(* Logix 5000 project; controller PLC_MCC1300_75F1 vendor 1 type 14 code 166 rev 32.11; software revision 32.04; part 69 of 83 *)
(* tags used below, declared in another part *)
   CM_LineToConveyorStacker_JS1 : CM_LineToConveyorStacker;
   GP_ScadaPlate : GP_ScadaPlate;
   M317 : MAC_Conveyor_Single;
   M317_ALM : MAC_Conveyor_ALM;
   M317_Data : UDT_Convoy_SL;
   M317_HMR : MAC_Conveyor_HMR;
   M317_HMW : MAC_Conveyor_HMW;
   M317_SpaceConv_Utilities : SpaceConv_Utilities;
   M317_TON_FrontSquarLeft_timeout : TIMER;
   M317_TON_FrontSquarRight_timeout : TIMER;
   M317_TON_LatSquarLeft_timeout : TIMER;
   M317_TON_LatSquarRight_timeout : TIMER;
   M317_TON_Synchro_timeout : TIMER;
   M317_xFrontLeftTimeout : BOOL;
   M317_xFrontRightTimeout : BOOL;
   M317_xLatLeftTimeout : BOOL;
   M317_xLatRightTimeout : BOOL;
   M317_xSensorTimeout : BOOL;
   M350Popup : MAC_Popup_ZC;
   M350Popup_ALM : MAC_Popup_ZC_ALM;
   M350Popup_HMR : MAC_Popup_ZC_HMR;
   M350Popup_HMW : MAC_Popup_ZC_HMW;
   O : INT[128];
   TMP_dHalfConveyorLength : DINT;
   TMP_xEnableZoneCleaning : BOOL;
   xAlwaysOFF : BOOL;
   xAlwaysON : BOOL;
   Z300_Conveyor : UDT_StandConv[29];
   Z300_LineTracking : UDT_LINE_TRACKING;
   Z301 : MAC_Zone_ML;
   Z402 : MAC_Zone;
   Z402_HMI_rgtPlateScada_Internal : HMI_LiteData[5,2,7];
(* MainProgram, continued *)

   // Command descent frontal squaring
   103: XIC(M317.ST_xManualMode)XIC(M317_HMW.rgxMan.17)XIC(M317.OUTPUT_xDescentSquaring_1)OTE(M317_HMR.rgxMan.17);
   // Commando conveyor M317 and conveyor stacker forward
   104: XIC(M317_HMW.rgxMan.25)XIC(M317.OUTPUT_xRun_M1)XIC(CM_LineToConveyorStacker_JS1.xManualCommandFwd)OTE(M317_HMR.rgxMan.25);
   // Commando conveyor M317 and conveyor stacker backward
   105: XIC(M317_HMW.rgxMan.26)XIC(M317.OUTPUT_xReverse_M1)XIC(CM_LineToConveyorStacker_JS1.xManualCommandBkw)OTE(M317_HMR.rgxMan.26);
   // Cleaning Enabled {x|x|x|x|O}
   106: XIC(M317.ST_xCleaningAccepted)[XIC(Z402.ST_xCleaningAccepted) ,XIO(TMP_xEnableZoneCleaning) ]OTE(M317_HMR.xCleaningEnabled);
   // Virtual door Enabled {x|x|x|x|O}
   107: XIC(M317.ST_xVirtualDoorEnabled)OTE(M317_HMR.xVirtualDoorEnabled);
   // Id plate presence
   108: XIC(M317.ST_xIdPlatePresence)OTE(M317_HMR.xIdPlatePresence);
   // Machine state M1
   109: XIC(xAlwaysON)[MOV(1,M317_HMR.dState1) ,XIC(M317.OUTPUT_xRun_M1) MOV(3,M317_HMR.dState1) ,XIC(M317.OUTPUT_xReverse_M1) MOV(4,M317_HMR.dState1) ,XIC(M317.ST_xMachineAlarm) MOV(7,M317_HMR.dState1) ];
   // Machine state M2
   110: XIC(xAlwaysON)[MOV(1,M317_HMR.dState2) ,XIC(M317.OUTPUT_xRun_M2) MOV(3,M317_HMR.dState2) ,XIC(M317.OUTPUT_xReverse_M2) MOV(4,M317_HMR.dState2) ,XIC(M317.ST_xMachineAlarm) MOV(7,M317_HMR.dState2) ];
   // Machine state M3
   111: XIC(xAlwaysON)[MOV(1,M317_HMR.dState3) ,XIC(M317.OUTPUT_xRun_M3) MOV(3,M317_HMR.dState3) ,XIC(M317.OUTPUT_xReverse_M3) MOV(4,M317_HMR.dState3) ,XIC(M317.ST_xMachineAlarm) MOV(7,M317_HMR.dState3) ];
   // Machine state M4
   112: XIC(xAlwaysON)[MOV(1,M317_HMR.dState4) ,XIC(M317.OUTPUT_xRun_M4) MOV(3,M317_HMR.dState4) ,XIC(M317.OUTPUT_xReverse_M4) MOV(4,M317_HMR.dState4) ,XIC(M317.ST_xMachineAlarm) MOV(7,M317_HMR.dState4) ];
   113: XIC(M317_SpaceConv_Utilities.O_xPlateSynchronized)OTE(M317.ST_xPlateSynchronized);
   114: XIC(M317.INPUT_xSyncroPhotocell_1)XIO(M317.ST_xIdPlatePresence)XIO(M317.ST_xPlatePresence)[TON(M317_TON_Synchro_timeout,?,?) ,[XIC(M317_TON_Synchro_timeout.DN) ,XIC(M317_xSensorTimeout) ] XIC(M317.INPUT_xSyncroPhotocell_1) OTE(M317_xSensorTimeout) ];
   115: XIC(M317.INPUT_xSquaringPhotocell_1)XIO(M317.ST_xIdPlatePresence)XIO(M317.ST_xPlatePresence)[TON(M317_TON_FrontSquarRight_timeout,?,?) ,[XIC(M317_TON_FrontSquarRight_timeout.DN) ,XIC(M317_xFrontRightTimeout) ] XIC(M317.INPUT_xSquaringPhotocell_1) OTE(M317_xFrontRightTimeout) ];
   116: XIC(M317.INPUT_xSquaringPhotocell_2)XIO(M317.ST_xIdPlatePresence)XIO(M317.ST_xPlatePresence)[TON(M317_TON_FrontSquarLeft_timeout,?,?) ,[XIC(M317_TON_FrontSquarLeft_timeout.DN) ,XIC(M317_xFrontLeftTimeout) ] XIC(M317.INPUT_xSquaringPhotocell_2) OTE(M317_xFrontLeftTimeout) ];
   117: XIC(M317.INPUT_xSquaringPhotocell_3)XIO(M317.ST_xIdPlatePresence)XIO(M317.ST_xPlatePresence)[TON(M317_TON_LatSquarRight_timeout,?,?) ,[XIC(M317_TON_LatSquarRight_timeout.DN) ,XIC(M317_xLatRightTimeout) ] XIC(M317.INPUT_xSquaringPhotocell_3) OTE(M317_xLatRightTimeout) ];
   118: XIC(M317.INPUT_xSquaringPhotocell_4)XIO(M317.ST_xIdPlatePresence)XIO(M317.ST_xPlatePresence)[TON(M317_TON_LatSquarLeft_timeout,?,?) ,[XIC(M317_TON_LatSquarLeft_timeout.DN) ,XIC(M317_xLatLeftTimeout) ] XIC(M317.INPUT_xSquaringPhotocell_4) OTE(M317_xLatLeftTimeout) ];
   // State Sensor
   119: XIC(xAlwaysON)[MOV(1,M317_HMR.dStateSensor5) ,XIC(M317_xSensorTimeout) MOV(7,M317_HMR.dStateSensor5) ];
   // State Sensor
   120: XIC(xAlwaysON)[MOV(1,M317_HMR.dStateSensor3) ,[XIC(M317_ALM.rgxStoppingFault[0].2) ,XIC(M317_ALM.rgxStoppingFault[0].3) ,XIC(M317_ALM.rgxWarning[0].25) ,XIC(M317_xFrontRightTimeout) ] MOV(7,M317_HMR.dStateSensor3) ];
   // State Sensor
   121: XIC(xAlwaysON)[MOV(1,M317_HMR.dStateSensor4) ,[XIC(M317_ALM.rgxStoppingFault[0].10) ,XIC(M317_ALM.rgxStoppingFault[0].11) ,XIC(M317_ALM.rgxWarning[0].25) ,XIC(M317_xFrontLeftTimeout) ] MOV(7,M317_HMR.dStateSensor4) ];
   // State Sensor
   122: XIC(xAlwaysON)[MOV(1,M317_HMR.dStateSensor1) ,[XIC(M317_ALM.rgxWarning[0].26) ,XIC(M317_xLatRightTimeout) ] MOV(7,M317_HMR.dStateSensor1) ];
   // State Sensor
   123: XIC(xAlwaysON)[MOV(1,M317_HMR.dStateSensor2) ,[XIC(M317_ALM.rgxWarning[0].26) ,XIC(M317_xLatLeftTimeout) ] MOV(7,M317_HMR.dStateSensor2) ];
   124: XIC(M317.ST_xIdPlatePresence)GP_ScadaPlate(GP_ScadaPlate,M317_Data,6,M317_SpaceConv_Utilities.O_dHeadPosition_cmm,M317_SpaceConv_Utilities.CONST_dConveyorWidth_cmm,M317_SpaceConv_Utilities.CONST_dConveyorLength_cmm,M317_SpaceConv_Utilities.ST_xLastModLoadBkw,M317_SpaceConv_Utilities.ST_xLastModUnloadBkw,1,0,Z402_HMI_rgtPlateScada_Internal);
END_ROUTINE

ROUTINE M350Popup_Faults   (* ladder *)
   // Reset faults
   0: XIC(Z301.ST_xAlarmOff)FLL(0,M350Popup_ALM,1);
   1: XIC(M350Popup.ST_xEnableControlError)[[XIC(M350Popup.OUTPUT_xPopupLifting) XIO(M350Popup.INPUT_xPopupHigh) ,XIO(M350Popup.OUTPUT_xPopupLifting) XIO(M350Popup.INPUT_xPopupLow) ,XIO(M350Popup.INPUT_xPopupHigh) XIO(M350Popup.INPUT_xPopupLow) ] XIO(M350Popup_ALM.rgxStoppingFault[0].0) TON(M350Popup.tmON_LiftingTimeOut,?,?) ,[XIC(M350Popup.tmON_LiftingTimeOut.DN) ,XIC(M350Popup.INPUT_xPopupHigh) XIC(M350Popup.INPUT_xPopupLow) ] OTL(M350Popup_ALM.rgxStoppingFault[0].0) ];
   2: XIC(xAlwaysOFF)XIC(M350Popup.ST_xEnableControlError)XIO(M350Popup.INPUT_xLiftingProtectionMotor)OTL(M350Popup_ALM.rgxFault[0].0);
   3: XIC(xAlwaysOFF)XIC(M350Popup.ST_xEnableControlError)[[XIC(M350Popup.OUTPUT_xPopupLifting) ,XIC(M350Popup.OUTPUT_xPopupDescent) ] XIO(M350Popup.INPUT_xLiftingFeedbackMotor) ,XIO(M350Popup.OUTPUT_xPopupLifting) XIO(M350Popup.OUTPUT_xPopupDescent) XIC(M350Popup.INPUT_xLiftingFeedbackMotor) ][TON(M350Popup.tmON_LiftingFeedbackTimeOut,?,?) ,XIC(M350Popup.tmON_LiftingFeedbackTimeOut.DN) OTL(M350Popup_ALM.rgxFault[0].1) ];
   4: XIC(xAlwaysOFF)XIC(M350Popup.ST_xEnableControlError)XIO(M350Popup.INPUT_xLiftingSafetySwitch)OTL(M350Popup_ALM.rgxFault[0].2);
   // Stopped machine fault
   5: [NEQ(M350Popup_ALM.rgxStoppingFault[0],0) ,NEQ(M350Popup_ALM.rgxStoppingFault_M[0],0) ]OTE(M350Popup.ST_xStopMachineFault);
   // Stopped next cycle fault
   6: [NEQ(M350Popup_ALM.rgxFault[0],0) ,NEQ(M350Popup_ALM.rgxFault_M[0],0) ]OTE(M350Popup.ST_xStopNextCycleFault);
   7: XIC(M350Popup.ST_xEnableControlError)XIC(M350Popup.ST_xOutputEnable)[XIC(M350Popup.PH_xRise) XIO(M350Popup.ST_xInitialConditionForRise) XIO(M350Popup.INPUT_xPopupHigh) ,XIC(M350Popup.PH_xDescend) XIO(M350Popup.ST_xInitialConditionForDescend) XIO(M350Popup.INPUT_xPopupLow) ]OTE(M350Popup.ST_xMachineWarning);
END_ROUTINE

ROUTINE M350Popup_Logic   (* ladder *)
   // #####_CONSTANTS_#####
   0: NOP();
   1: XIC(xAlwaysON)OTE(M350Popup.ST_xTunnelType);
   2: DIV(Z300_LineTracking.rgtTrkConv[21].dLengthConveyor,2,TMP_dHalfConveyorLength);
   3: MOV(Z300_LineTracking.rgtTrkConv[21].dStartPosition_cmm,M350Popup.AUX_dStartPosition_cmm)MOV(Z300_LineTracking.rgtTrkConv[21].dEndPosition_cmm,M350Popup.AUX_dEndPosition_cmm)MOV(1500,M350Popup.AUX_dReactionTime_ms)MOV(200000,M350Popup.AUX_dWindowSearch_cmm)MOV(Z300_Conveyor[21].AUX_rgdCurrentSpeed_mm_min[0],M350Popup.AUX_dSpeedConveyor_mm_min);
   // #####_MATCH_#####
   4: NOP();
   5: XIC(Z301.ST_xEnableControlError)OTE(M350Popup.ST_xEnableControlError);
   // #####_ALARMS_#####
   6: NOP();
   7: JSR(M350Popup_Faults,0);
   // #####_HMI_LOGICS_#####
   8: NOP();
   9: XIC(xAlwaysON)OTE(M350Popup.ST_xExternalConditionToRise);
   10: XIC(xAlwaysON)OTE(M350Popup.ST_xExternalConditionToDescend);
   // #####_STATUSES_#####
   11: NOP();
   12: [XIC(M350Popup.ST_xStopMachineFault) ,XIC(M350Popup.ST_xStopNextCycleFault) ]OTE(M350Popup.ST_xMachineAlarm);
   13: [XIO(M350Popup.ST_xPhasesInProgress) ,XIO(M350Popup.ST_xOutputEnable) ]OTE(M350Popup.ST_xConditionOKForStopCycle);
   14: XIC(Z301.ST_xCycleON)XIO(M350Popup.ST_xManualMode)XIO(M350Popup.ST_xMachineAlarm)OTE(M350Popup.ST_xOutputEnable);
   15: XIC(Z301.ST_xCycleON)XIC(M350Popup.ST_xOutputEnable)XIO(M350Popup.ST_xPhasesInProgress)XIO(M350Popup.INPUT_xPopupHigh)XIO(M350Popup.ST_xCleaningAccepted)OTE(M350Popup.ST_xInitialConditionForRise);
   16: XIC(Z301.ST_xCycleON)XIC(M350Popup.ST_xOutputEnable)XIO(M350Popup.ST_xPhasesInProgress)XIO(M350Popup.INPUT_xPopupLow)XIO(M350Popup.ST_xCleaningAccepted)OTE(M350Popup.ST_xInitialConditionForDescend);
   17: [XIC(M350Popup_HMW.xEnableDisableManualCommand) XIC(xAlwaysOFF) ,XIC(Z300_Conveyor[21].ST_xManualCmdEnabled) ]XIC(M350Popup.ST_xConditionOKForStopCycle)OTE(M350Popup.ST_xManualMode);
   18: XIO(M350Popup.ST_xManualMode)MOV(0,M350Popup_HMW.rgxMan);
   // #####_PHASES_&_LOGICS_#####
   19: NOP();
   20: XIC(xAlwaysON)OTE(M350Popup.ST_xCleaningConditionOK);
   21: [XIC(M350Popup_HMW.xLocalCleaningRequest) XIC(xAlwaysOFF) ,XIC(Z300_Conveyor[21].ST_xCleaningEnabled) XIC(M350Popup.INPUT_xPopupLow) ][XIC(M350Popup.ST_xCleaningConditionOK) ,XIC(M350Popup.ST_xCleaningAccepted) ]OTE(M350Popup.ST_xCleaningAccepted);
   22: XIC(M350Popup.ST_xInitialConditionForRise)XIC(M350Popup.ST_xExternalConditionToRise)XIC(M350Popup.ST_xRequestRise)XIO(M350Popup.PH_xRise)OTL(M350Popup.PH_xRise);
   23: XIC(M350Popup.PH_xRise)XIC(M350Popup.INPUT_xPopupHigh)XIO(M350Popup.INPUT_xPopupLow)[XIC(M350Popup.INPUT_xPopupHigh) OTU(M350Popup.PH_xRise) ,OTE(M350Popup.PH_xEndRise) ];
   24: XIC(M350Popup.ST_xInitialConditionForDescend)XIC(M350Popup.ST_xExternalConditionToDescend)XIC(M350Popup.ST_xRequestDescend)XIO(M350Popup.PH_xDescend)OTL(M350Popup.PH_xDescend);
   25: XIC(M350Popup.PH_xDescend)XIC(M350Popup.INPUT_xPopupLow)XIO(M350Popup.INPUT_xPopupHigh)[OTU(M350Popup.PH_xDescend) ,OTE(M350Popup.PH_xEndDescend) ];
   26: [XIC(M350Popup.PH_xRise) ,XIC(M350Popup.PH_xEndRise) ,XIC(M350Popup.PH_xDescend) ,XIC(M350Popup.PH_xEndDescend) ]OTE(M350Popup.ST_xPhasesInProgress);
   27: [XIC(M350Popup.PH_xEndDescend) ,XIC(M350Popup.INPUT_xPopupLow) ]OTU(M350Popup.ST_xPlatePresence);
   28: XIO(M350Popup.ST_xPhasesInProgress)[XIC(M350Popup.INPUT_xPopupLow) XIO(M350Popup.INPUT_xPopupHigh) ,XIC(M350Popup.ST_xTunnelType) XIC(M350Popup.INPUT_xPopupHigh) XIO(M350Popup.INPUT_xPopupLow) ]OTE(M350Popup.ST_xOutOfEncumbrance);
   29: XIO(M350Popup.ST_xPhasesInProgress)XIO(M350Popup.ST_xPlatePresence)XIO(M350Popup.INPUT_xPopupHigh)XIC(M350Popup.INPUT_xPopupLow)OTE(M350Popup.ST_xConditionToReceiveGlass);
   30: XIO(M350Popup.ST_xPhasesInProgress)XIC(M350Popup.INPUT_xPopupHigh)XIO(M350Popup.INPUT_xPopupLow)OTE(M350Popup.ST_xConditionForUpperConveyor);
   // #####_EXTERNAL_DEVICE_#####
   31: NOP();
   // #####_HMI_STATUSES_#####
   32: NOP();
   33: XIC(M350Popup.INPUT_xPopupHigh)OTE(M350Popup_HMR.xHighPosition);
   34: XIC(M350Popup.INPUT_xPopupLow)OTE(M350Popup_HMR.xLowPosition);
   35: [MOV(1,M350Popup_HMR.rgdState) ,[XIC(M350Popup.OUTPUT_xPopupLifting) ,XIC(M350Popup.OUTPUT_xPopupDescent) ] MOV(3,M350Popup_HMR.rgdState) ,XIC(M350Popup.ST_xMachineWarning) MOV(5,M350Popup_HMR.rgdState) ,XIC(M350Popup.ST_xMachineAlarm) MOV(7,M350Popup_HMR.rgdState) ];
   36: XIC(M350Popup.ST_xCleaningAccepted)OTE(M350Popup_HMR.xPopUpCleaningEnabled);
   37: XIC(M350Popup.ST_xManualMode)XIC(M350Popup_HMW.rgxMan.0)XIC(M350Popup.OUTPUT_xPopupLifting)OTE(M350Popup_HMR.rgxMan.0);
   38: XIC(M350Popup.ST_xManualMode)XIC(M350Popup_HMW.rgxMan.1)XIC(M350Popup.OUTPUT_xPopupDescent)OTE(M350Popup_HMR.rgxMan.1);
   39: XIC(M350Popup.ST_xManualMode)XIC(M350Popup_HMW.rgxMan.8)XIC(M350Popup.OUTPUT_xRun)OTE(M350Popup_HMR.rgxMan.8);
   40: XIC(M350Popup.ST_xManualMode)XIC(M350Popup_HMW.rgxMan.9)XIC(M350Popup.OUTPUT_xReverse)OTE(M350Popup_HMR.rgxMan.9);
END_ROUTINE
